(* Logix 5000 project; controller PLC_MCC1300_75F1 vendor 1 type 14 code 166 rev 32.11; software revision 32.04; part 12 of 83 *)
(* tags used below, declared in another part *)
   M302SpeedUp : MAC_SpeedUp;
   TMP_d : DINT;
   TMP_xPositioning : BOOL;
   TMP_xReverse : BOOL;
   TMP_xRun : BOOL;
   xAlwaysOFF : BOOL;
   Z300_Conveyor : UDT_StandConv[29];
   Z300_Conveyor_Conf : UDT_Conveyor_Config[29];
   Z300_Conveyor_HMW : MAC_Conveyor_ZC_HMW[29];
   Z300_Conveyor_IN_MOTION : MAC_Conveyor_ZC_IN_MOTION[29];
   Z301_HMR : MAC_Zone_ML_HMR;
(* CommandLogic, continued *)

ROUTINE M302M2_Conveyor_Output   (* ladder *)
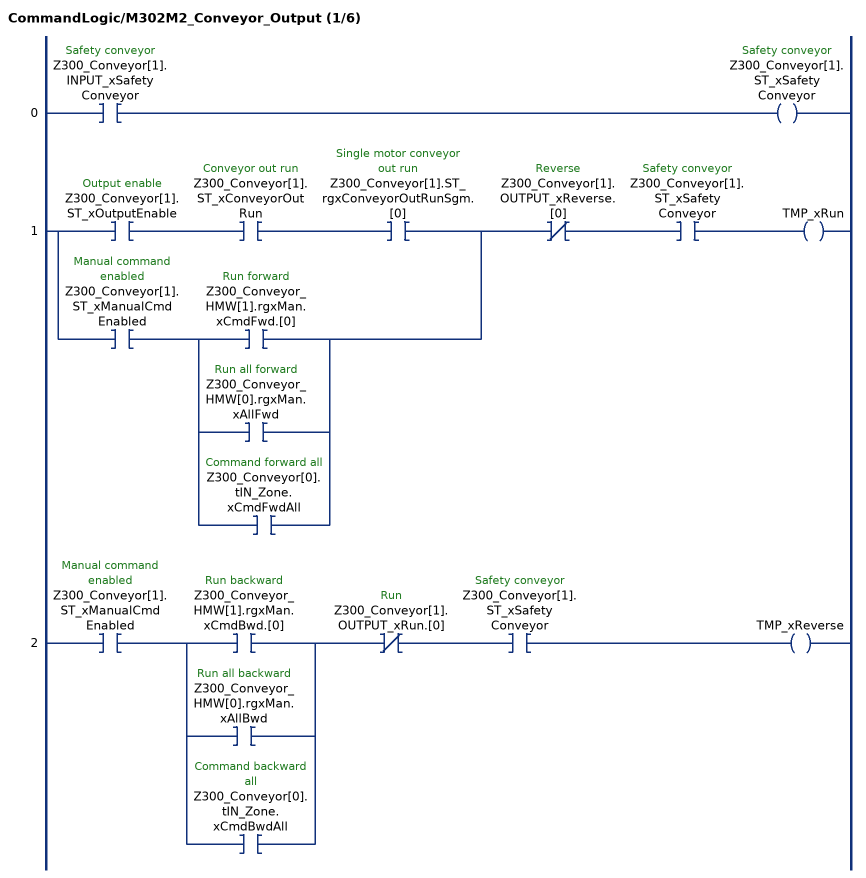
   0: XIC(Z300_Conveyor[1].INPUT_xSafetyConveyor)OTE(Z300_Conveyor[1].ST_xSafetyConveyor);
   1: [XIC(Z300_Conveyor[1].ST_xOutputEnable) XIC(Z300_Conveyor[1].ST_xConveyorOutRun) XIC(Z300_Conveyor[1].ST_rgxConveyorOutRunSgm.[0]) ,XIC(Z300_Conveyor[1].ST_xManualCmdEnabled) [XIC(Z300_Conveyor_HMW[1].rgxMan.xCmdFwd.[0]) ,XIC(Z300_Conveyor_HMW[0].rgxMan.xAllFwd) ,XIC(Z300_Conveyor[0].tIN_Zone.xCmdFwdAll) ] ]XIO(Z300_Conveyor[1].OUTPUT_xReverse.[0])XIC(Z300_Conveyor[1].ST_xSafetyConveyor)OTE(TMP_xRun);
   2: XIC(Z300_Conveyor[1].ST_xManualCmdEnabled)[XIC(Z300_Conveyor_HMW[1].rgxMan.xCmdBwd.[0]) ,XIC(Z300_Conveyor_HMW[0].rgxMan.xAllBwd) ,XIC(Z300_Conveyor[0].tIN_Zone.xCmdBwdAll) ]XIO(Z300_Conveyor[1].OUTPUT_xRun.[0])XIC(Z300_Conveyor[1].ST_xSafetyConveyor)OTE(TMP_xReverse);
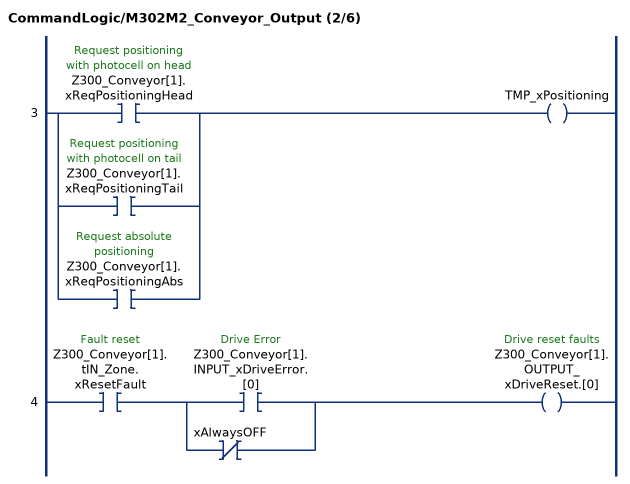
   3: [XIC(Z300_Conveyor[1].xReqPositioningHead) ,XIC(Z300_Conveyor[1].xReqPositioningTail) ,XIC(Z300_Conveyor[1].xReqPositioningAbs) ]OTE(TMP_xPositioning);
   4: XIC(Z300_Conveyor[1].tIN_Zone.xResetFault)[XIC(Z300_Conveyor[1].INPUT_xDriveError.[0]) ,XIO(xAlwaysOFF) ]OTE(Z300_Conveyor[1].OUTPUT_xDriveReset.[0]);
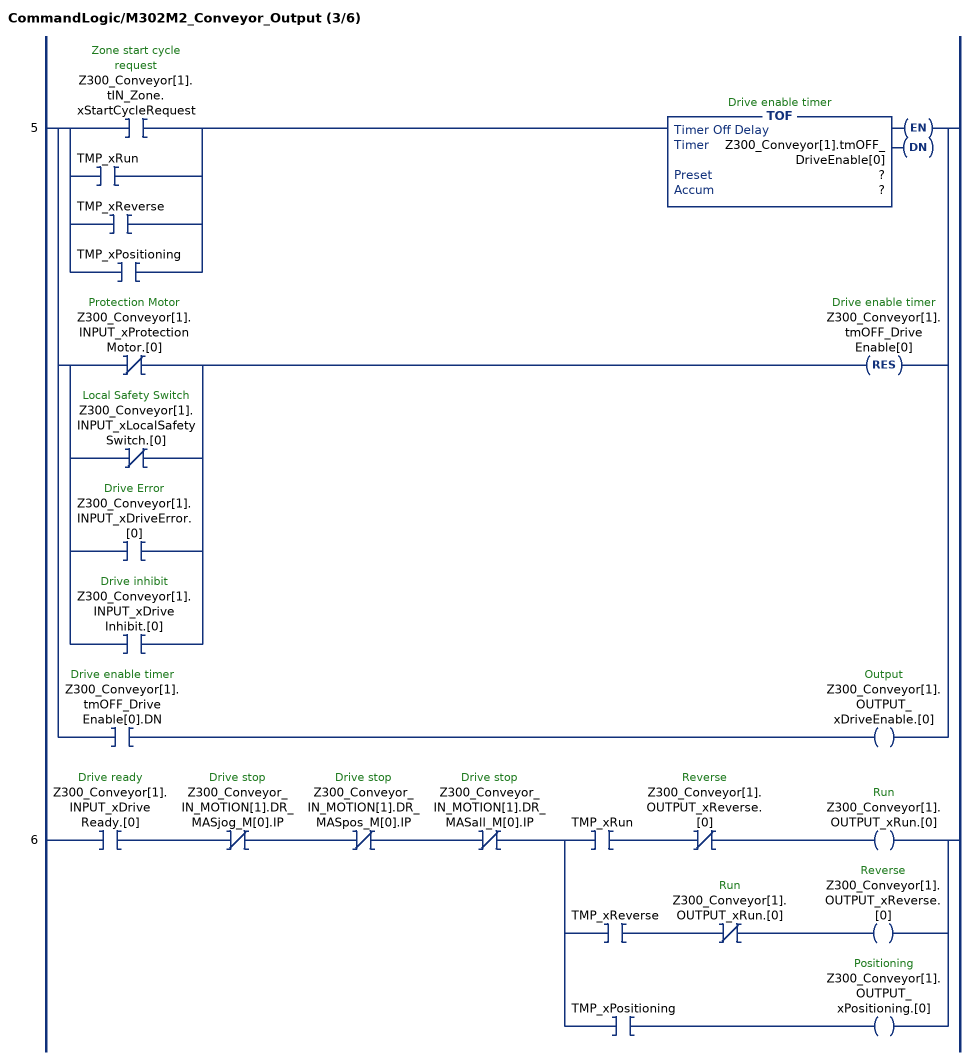
   5: [[XIC(Z300_Conveyor[1].tIN_Zone.xStartCycleRequest) ,XIC(TMP_xRun) ,XIC(TMP_xReverse) ,XIC(TMP_xPositioning) ] TOF(Z300_Conveyor[1].tmOFF_DriveEnable[0],?,?) ,[XIO(Z300_Conveyor[1].INPUT_xProtectionMotor.[0]) ,XIO(Z300_Conveyor[1].INPUT_xLocalSafetySwitch.[0]) ,XIC(Z300_Conveyor[1].INPUT_xDriveError.[0]) ,XIC(Z300_Conveyor[1].INPUT_xDriveInhibit.[0]) ] RES(Z300_Conveyor[1].tmOFF_DriveEnable[0]) ,XIC(Z300_Conveyor[1].tmOFF_DriveEnable[0].DN) OTE(Z300_Conveyor[1].OUTPUT_xDriveEnable.[0]) ];
   6: XIC(Z300_Conveyor[1].INPUT_xDriveReady.[0])XIO(Z300_Conveyor_IN_MOTION[1].DR_MASjog_M[0].IP)XIO(Z300_Conveyor_IN_MOTION[1].DR_MASpos_M[0].IP)XIO(Z300_Conveyor_IN_MOTION[1].DR_MASall_M[0].IP)[XIC(TMP_xRun) XIO(Z300_Conveyor[1].OUTPUT_xReverse.[0]) OTE(Z300_Conveyor[1].OUTPUT_xRun.[0]) ,XIC(TMP_xReverse) XIO(Z300_Conveyor[1].OUTPUT_xRun.[0]) OTE(Z300_Conveyor[1].OUTPUT_xReverse.[0]) ,XIC(TMP_xPositioning) OTE(Z300_Conveyor[1].OUTPUT_xPositioning.[0]) ];
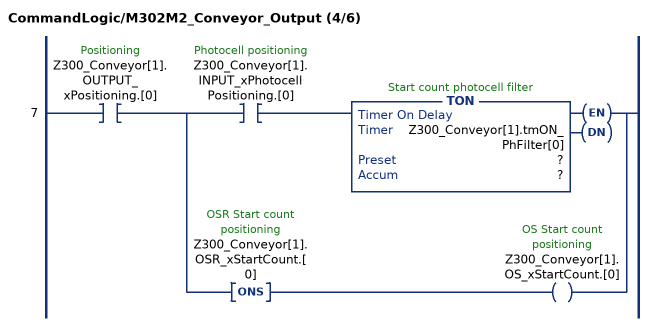
   7: XIC(Z300_Conveyor[1].OUTPUT_xPositioning.[0])[XIC(Z300_Conveyor[1].INPUT_xPhotocellPositioning.[0]) TON(Z300_Conveyor[1].tmON_PhFilter[0],?,?) ,ONS(Z300_Conveyor[1].OSR_xStartCount.[0]) OTE(Z300_Conveyor[1].OS_xStartCount.[0]) ];
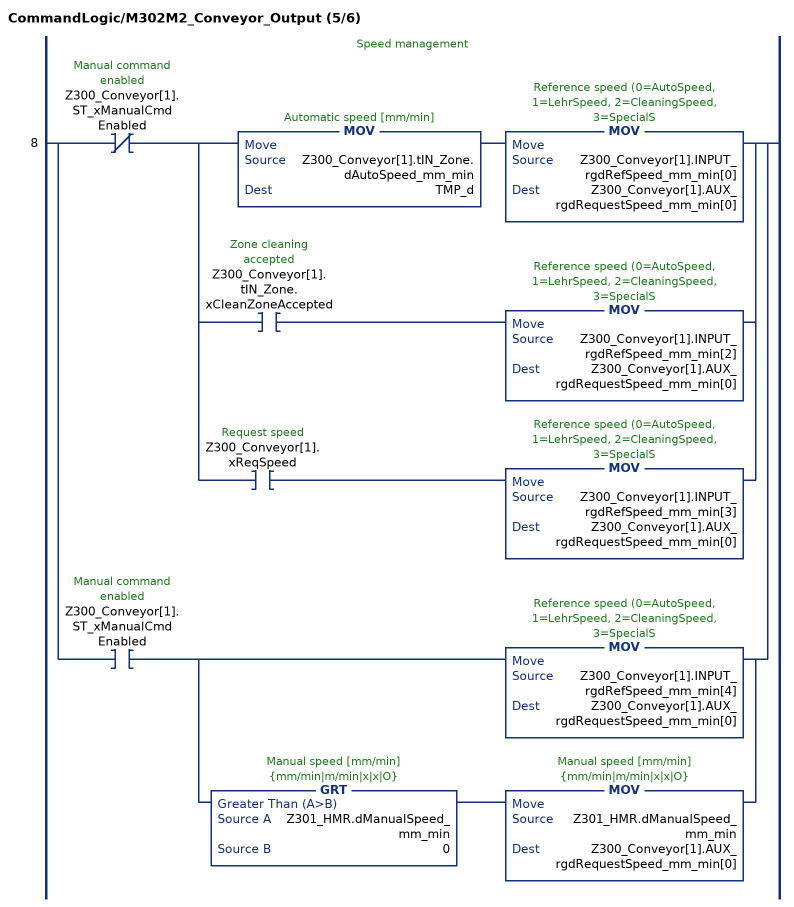
   // Speed management
   8: [XIO(Z300_Conveyor[1].ST_xManualCmdEnabled) [MOV(Z300_Conveyor[1].tIN_Zone.dAutoSpeed_mm_min,TMP_d) MOV(Z300_Conveyor[1].INPUT_rgdRefSpeed_mm_min[0],Z300_Conveyor[1].AUX_rgdRequestSpeed_mm_min[0]) ,XIC(Z300_Conveyor[1].tIN_Zone.xCleanZoneAccepted) MOV(Z300_Conveyor[1].INPUT_rgdRefSpeed_mm_min[2],Z300_Conveyor[1].AUX_rgdRequestSpeed_mm_min[0]) ,XIC(Z300_Conveyor[1].xReqSpeed) MOV(Z300_Conveyor[1].INPUT_rgdRefSpeed_mm_min[3],Z300_Conveyor[1].AUX_rgdRequestSpeed_mm_min[0]) ] ,XIC(Z300_Conveyor[1].ST_xManualCmdEnabled) [MOV(Z300_Conveyor[1].INPUT_rgdRefSpeed_mm_min[4],Z300_Conveyor[1].AUX_rgdRequestSpeed_mm_min[0]) ,GRT(Z301_HMR.dManualSpeed_mm_min,0) MOV(Z301_HMR.dManualSpeed_mm_min,Z300_Conveyor[1].AUX_rgdRequestSpeed_mm_min[0]) ] ];
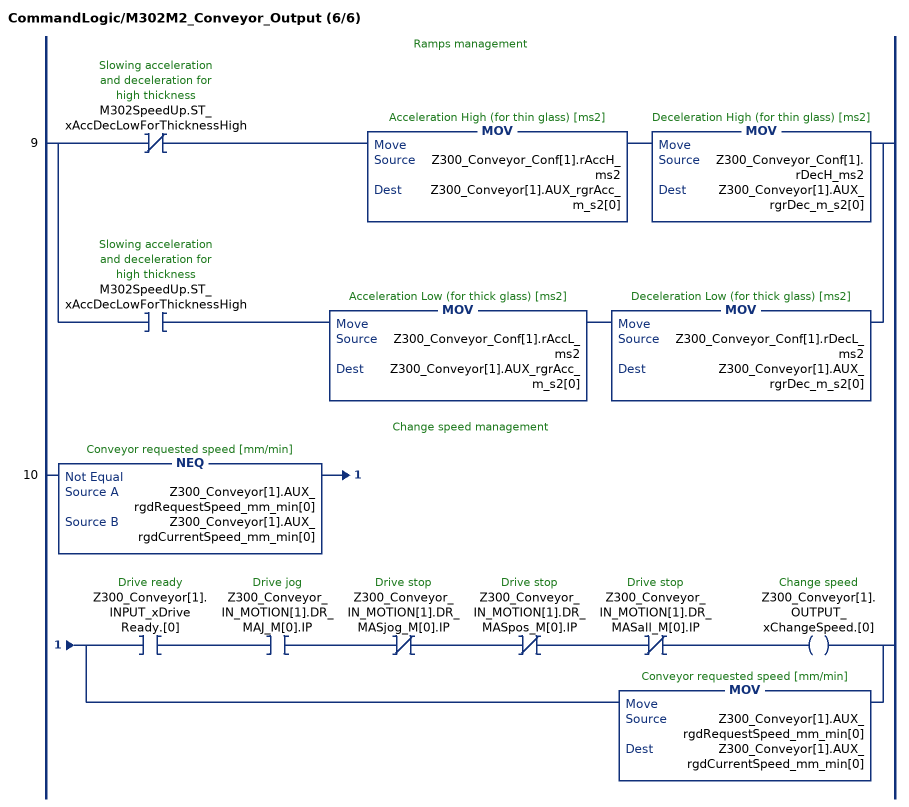
   // Ramps management
   9: [XIO(M302SpeedUp.ST_xAccDecLowForThicknessHigh) MOV(Z300_Conveyor_Conf[1].rAccH_ms2,Z300_Conveyor[1].AUX_rgrAcc_m_s2[0]) MOV(Z300_Conveyor_Conf[1].rDecH_ms2,Z300_Conveyor[1].AUX_rgrDec_m_s2[0]) ,XIC(M302SpeedUp.ST_xAccDecLowForThicknessHigh) MOV(Z300_Conveyor_Conf[1].rAccL_ms2,Z300_Conveyor[1].AUX_rgrAcc_m_s2[0]) MOV(Z300_Conveyor_Conf[1].rDecL_ms2,Z300_Conveyor[1].AUX_rgrDec_m_s2[0]) ];
   // Change speed management
   10: NEQ(Z300_Conveyor[1].AUX_rgdRequestSpeed_mm_min[0],Z300_Conveyor[1].AUX_rgdCurrentSpeed_mm_min[0])[XIC(Z300_Conveyor[1].INPUT_xDriveReady.[0]) XIC(Z300_Conveyor_IN_MOTION[1].DR_MAJ_M[0].IP) XIO(Z300_Conveyor_IN_MOTION[1].DR_MASjog_M[0].IP) XIO(Z300_Conveyor_IN_MOTION[1].DR_MASpos_M[0].IP) XIO(Z300_Conveyor_IN_MOTION[1].DR_MASall_M[0].IP) OTE(Z300_Conveyor[1].OUTPUT_xChangeSpeed.[0]) ,MOV(Z300_Conveyor[1].AUX_rgdRequestSpeed_mm_min[0],Z300_Conveyor[1].AUX_rgdCurrentSpeed_mm_min[0]) ];
END_ROUTINE

ROUTINE M302M3_Conveyor_Output   (* ladder *)
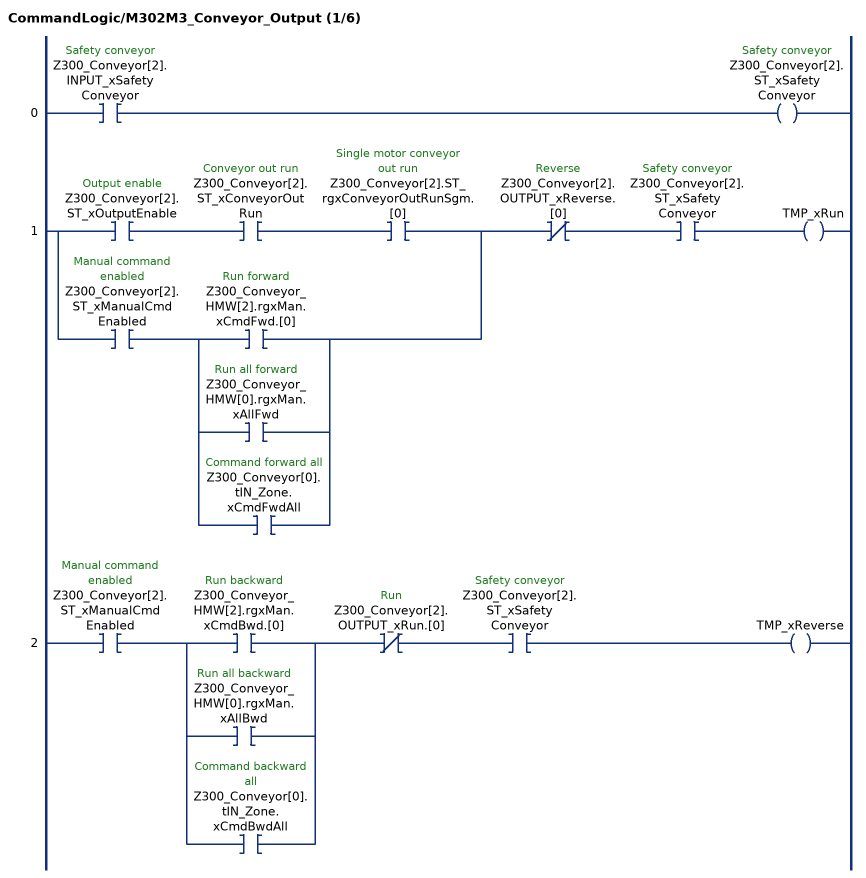
   0: XIC(Z300_Conveyor[2].INPUT_xSafetyConveyor)OTE(Z300_Conveyor[2].ST_xSafetyConveyor);
   1: [XIC(Z300_Conveyor[2].ST_xOutputEnable) XIC(Z300_Conveyor[2].ST_xConveyorOutRun) XIC(Z300_Conveyor[2].ST_rgxConveyorOutRunSgm.[0]) ,XIC(Z300_Conveyor[2].ST_xManualCmdEnabled) [XIC(Z300_Conveyor_HMW[2].rgxMan.xCmdFwd.[0]) ,XIC(Z300_Conveyor_HMW[0].rgxMan.xAllFwd) ,XIC(Z300_Conveyor[0].tIN_Zone.xCmdFwdAll) ] ]XIO(Z300_Conveyor[2].OUTPUT_xReverse.[0])XIC(Z300_Conveyor[2].ST_xSafetyConveyor)OTE(TMP_xRun);
   2: XIC(Z300_Conveyor[2].ST_xManualCmdEnabled)[XIC(Z300_Conveyor_HMW[2].rgxMan.xCmdBwd.[0]) ,XIC(Z300_Conveyor_HMW[0].rgxMan.xAllBwd) ,XIC(Z300_Conveyor[0].tIN_Zone.xCmdBwdAll) ]XIO(Z300_Conveyor[2].OUTPUT_xRun.[0])XIC(Z300_Conveyor[2].ST_xSafetyConveyor)OTE(TMP_xReverse);
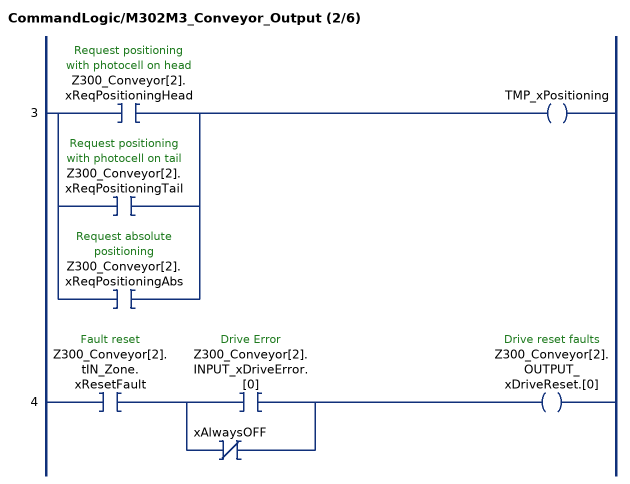
   3: [XIC(Z300_Conveyor[2].xReqPositioningHead) ,XIC(Z300_Conveyor[2].xReqPositioningTail) ,XIC(Z300_Conveyor[2].xReqPositioningAbs) ]OTE(TMP_xPositioning);
   4: XIC(Z300_Conveyor[2].tIN_Zone.xResetFault)[XIC(Z300_Conveyor[2].INPUT_xDriveError.[0]) ,XIO(xAlwaysOFF) ]OTE(Z300_Conveyor[2].OUTPUT_xDriveReset.[0]);
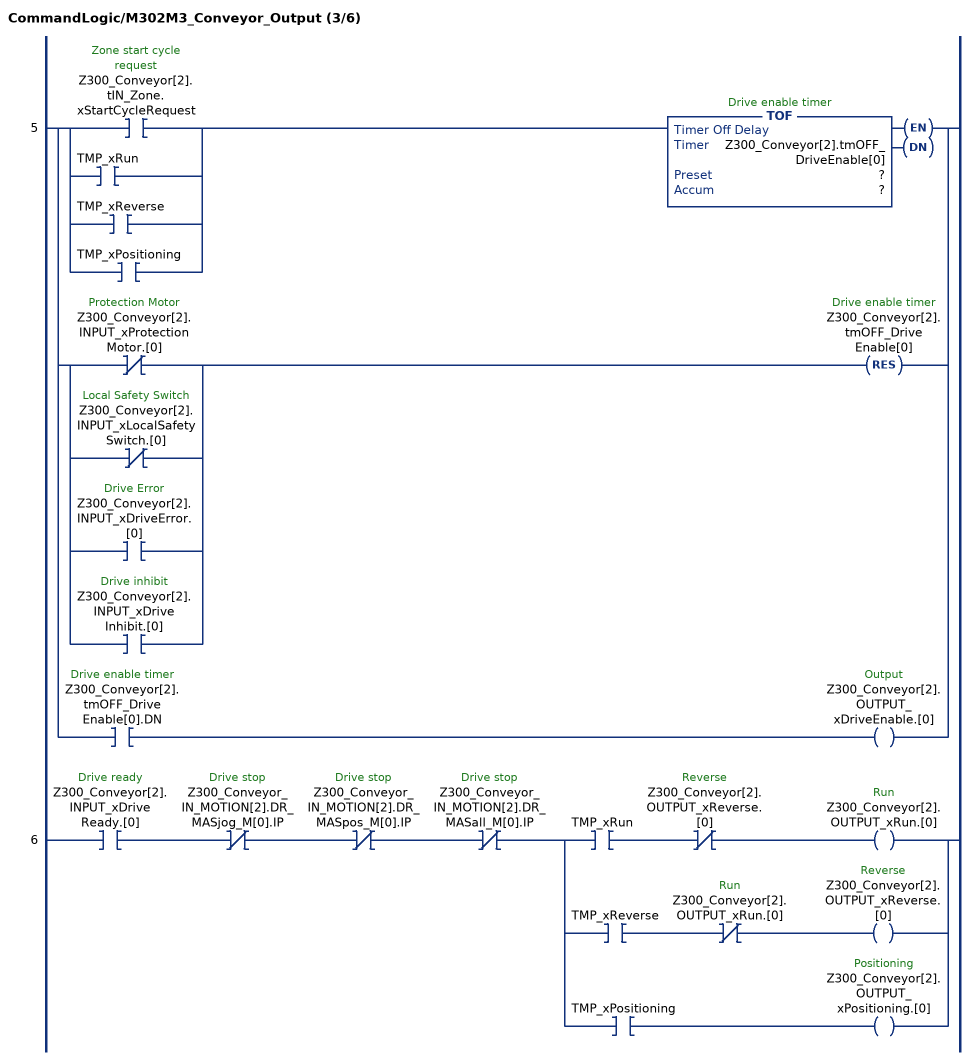
   5: [[XIC(Z300_Conveyor[2].tIN_Zone.xStartCycleRequest) ,XIC(TMP_xRun) ,XIC(TMP_xReverse) ,XIC(TMP_xPositioning) ] TOF(Z300_Conveyor[2].tmOFF_DriveEnable[0],?,?) ,[XIO(Z300_Conveyor[2].INPUT_xProtectionMotor.[0]) ,XIO(Z300_Conveyor[2].INPUT_xLocalSafetySwitch.[0]) ,XIC(Z300_Conveyor[2].INPUT_xDriveError.[0]) ,XIC(Z300_Conveyor[2].INPUT_xDriveInhibit.[0]) ] RES(Z300_Conveyor[2].tmOFF_DriveEnable[0]) ,XIC(Z300_Conveyor[2].tmOFF_DriveEnable[0].DN) OTE(Z300_Conveyor[2].OUTPUT_xDriveEnable.[0]) ];
   6: XIC(Z300_Conveyor[2].INPUT_xDriveReady.[0])XIO(Z300_Conveyor_IN_MOTION[2].DR_MASjog_M[0].IP)XIO(Z300_Conveyor_IN_MOTION[2].DR_MASpos_M[0].IP)XIO(Z300_Conveyor_IN_MOTION[2].DR_MASall_M[0].IP)[XIC(TMP_xRun) XIO(Z300_Conveyor[2].OUTPUT_xReverse.[0]) OTE(Z300_Conveyor[2].OUTPUT_xRun.[0]) ,XIC(TMP_xReverse) XIO(Z300_Conveyor[2].OUTPUT_xRun.[0]) OTE(Z300_Conveyor[2].OUTPUT_xReverse.[0]) ,XIC(TMP_xPositioning) OTE(Z300_Conveyor[2].OUTPUT_xPositioning.[0]) ];
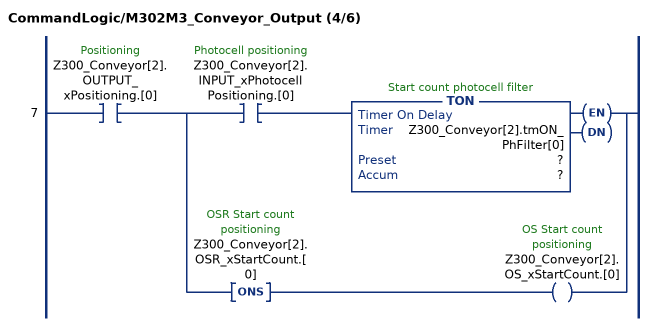
   7: XIC(Z300_Conveyor[2].OUTPUT_xPositioning.[0])[XIC(Z300_Conveyor[2].INPUT_xPhotocellPositioning.[0]) TON(Z300_Conveyor[2].tmON_PhFilter[0],?,?) ,ONS(Z300_Conveyor[2].OSR_xStartCount.[0]) OTE(Z300_Conveyor[2].OS_xStartCount.[0]) ];
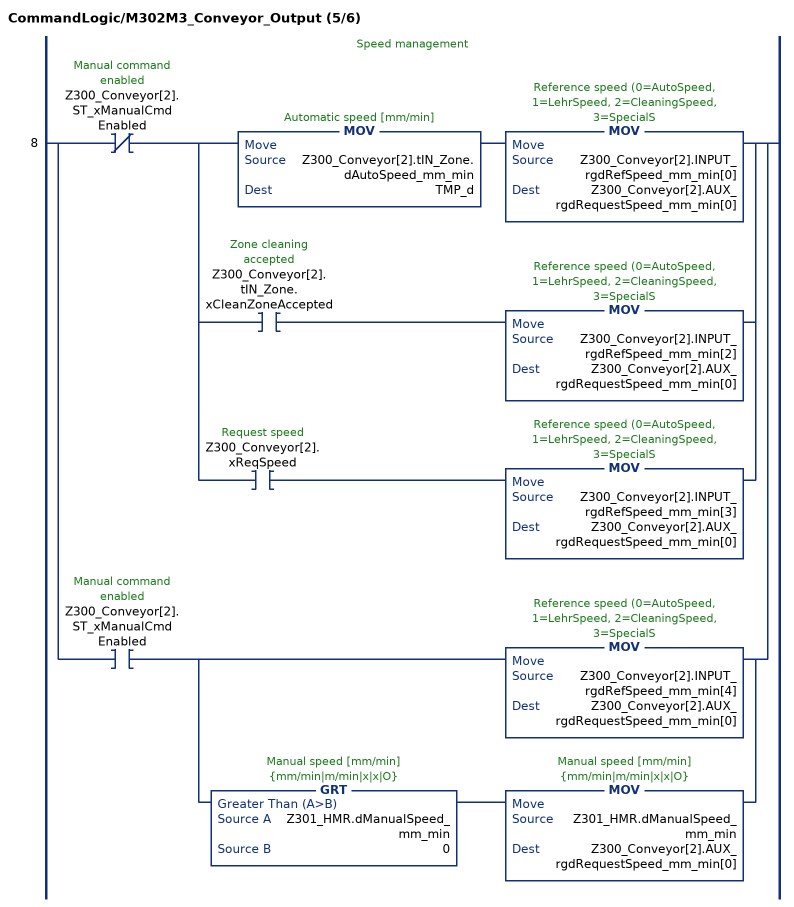
   // Speed management
   8: [XIO(Z300_Conveyor[2].ST_xManualCmdEnabled) [MOV(Z300_Conveyor[2].tIN_Zone.dAutoSpeed_mm_min,TMP_d) MOV(Z300_Conveyor[2].INPUT_rgdRefSpeed_mm_min[0],Z300_Conveyor[2].AUX_rgdRequestSpeed_mm_min[0]) ,XIC(Z300_Conveyor[2].tIN_Zone.xCleanZoneAccepted) MOV(Z300_Conveyor[2].INPUT_rgdRefSpeed_mm_min[2],Z300_Conveyor[2].AUX_rgdRequestSpeed_mm_min[0]) ,XIC(Z300_Conveyor[2].xReqSpeed) MOV(Z300_Conveyor[2].INPUT_rgdRefSpeed_mm_min[3],Z300_Conveyor[2].AUX_rgdRequestSpeed_mm_min[0]) ] ,XIC(Z300_Conveyor[2].ST_xManualCmdEnabled) [MOV(Z300_Conveyor[2].INPUT_rgdRefSpeed_mm_min[4],Z300_Conveyor[2].AUX_rgdRequestSpeed_mm_min[0]) ,GRT(Z301_HMR.dManualSpeed_mm_min,0) MOV(Z301_HMR.dManualSpeed_mm_min,Z300_Conveyor[2].AUX_rgdRequestSpeed_mm_min[0]) ] ];
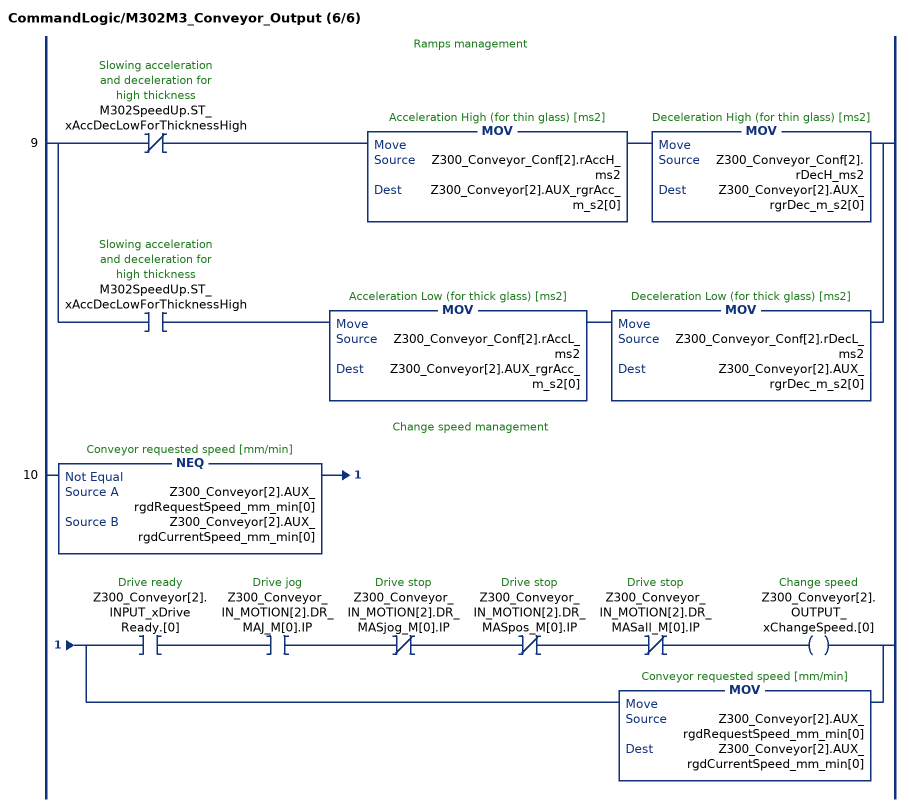
   // Ramps management
   9: [XIO(M302SpeedUp.ST_xAccDecLowForThicknessHigh) MOV(Z300_Conveyor_Conf[2].rAccH_ms2,Z300_Conveyor[2].AUX_rgrAcc_m_s2[0]) MOV(Z300_Conveyor_Conf[2].rDecH_ms2,Z300_Conveyor[2].AUX_rgrDec_m_s2[0]) ,XIC(M302SpeedUp.ST_xAccDecLowForThicknessHigh) MOV(Z300_Conveyor_Conf[2].rAccL_ms2,Z300_Conveyor[2].AUX_rgrAcc_m_s2[0]) MOV(Z300_Conveyor_Conf[2].rDecL_ms2,Z300_Conveyor[2].AUX_rgrDec_m_s2[0]) ];
   // Change speed management
   10: NEQ(Z300_Conveyor[2].AUX_rgdRequestSpeed_mm_min[0],Z300_Conveyor[2].AUX_rgdCurrentSpeed_mm_min[0])[XIC(Z300_Conveyor[2].INPUT_xDriveReady.[0]) XIC(Z300_Conveyor_IN_MOTION[2].DR_MAJ_M[0].IP) XIO(Z300_Conveyor_IN_MOTION[2].DR_MASjog_M[0].IP) XIO(Z300_Conveyor_IN_MOTION[2].DR_MASpos_M[0].IP) XIO(Z300_Conveyor_IN_MOTION[2].DR_MASall_M[0].IP) OTE(Z300_Conveyor[2].OUTPUT_xChangeSpeed.[0]) ,MOV(Z300_Conveyor[2].AUX_rgdRequestSpeed_mm_min[0],Z300_Conveyor[2].AUX_rgdCurrentSpeed_mm_min[0]) ];
END_ROUTINE

ROUTINE M302M4_Conveyor_Output   (* ladder *)
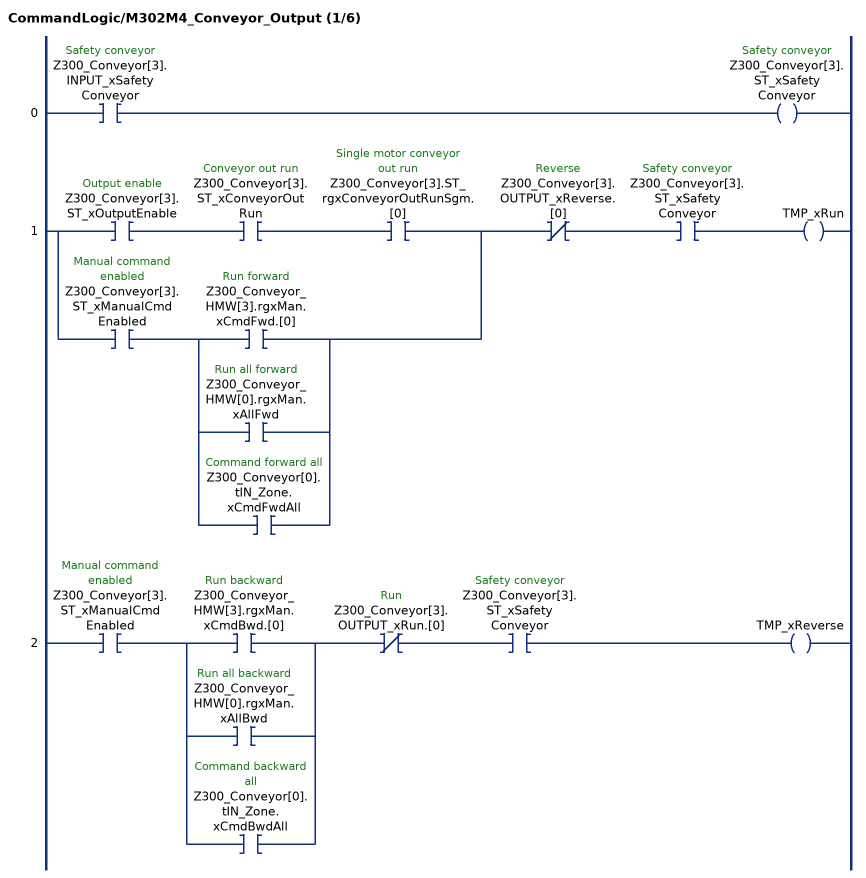
   0: XIC(Z300_Conveyor[3].INPUT_xSafetyConveyor)OTE(Z300_Conveyor[3].ST_xSafetyConveyor);
   1: [XIC(Z300_Conveyor[3].ST_xOutputEnable) XIC(Z300_Conveyor[3].ST_xConveyorOutRun) XIC(Z300_Conveyor[3].ST_rgxConveyorOutRunSgm.[0]) ,XIC(Z300_Conveyor[3].ST_xManualCmdEnabled) [XIC(Z300_Conveyor_HMW[3].rgxMan.xCmdFwd.[0]) ,XIC(Z300_Conveyor_HMW[0].rgxMan.xAllFwd) ,XIC(Z300_Conveyor[0].tIN_Zone.xCmdFwdAll) ] ]XIO(Z300_Conveyor[3].OUTPUT_xReverse.[0])XIC(Z300_Conveyor[3].ST_xSafetyConveyor)OTE(TMP_xRun);
   2: XIC(Z300_Conveyor[3].ST_xManualCmdEnabled)[XIC(Z300_Conveyor_HMW[3].rgxMan.xCmdBwd.[0]) ,XIC(Z300_Conveyor_HMW[0].rgxMan.xAllBwd) ,XIC(Z300_Conveyor[0].tIN_Zone.xCmdBwdAll) ]XIO(Z300_Conveyor[3].OUTPUT_xRun.[0])XIC(Z300_Conveyor[3].ST_xSafetyConveyor)OTE(TMP_xReverse);
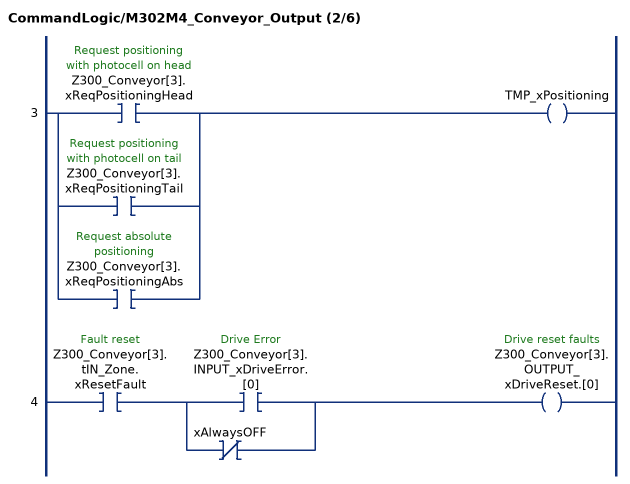
   3: [XIC(Z300_Conveyor[3].xReqPositioningHead) ,XIC(Z300_Conveyor[3].xReqPositioningTail) ,XIC(Z300_Conveyor[3].xReqPositioningAbs) ]OTE(TMP_xPositioning);
   4: XIC(Z300_Conveyor[3].tIN_Zone.xResetFault)[XIC(Z300_Conveyor[3].INPUT_xDriveError.[0]) ,XIO(xAlwaysOFF) ]OTE(Z300_Conveyor[3].OUTPUT_xDriveReset.[0]);
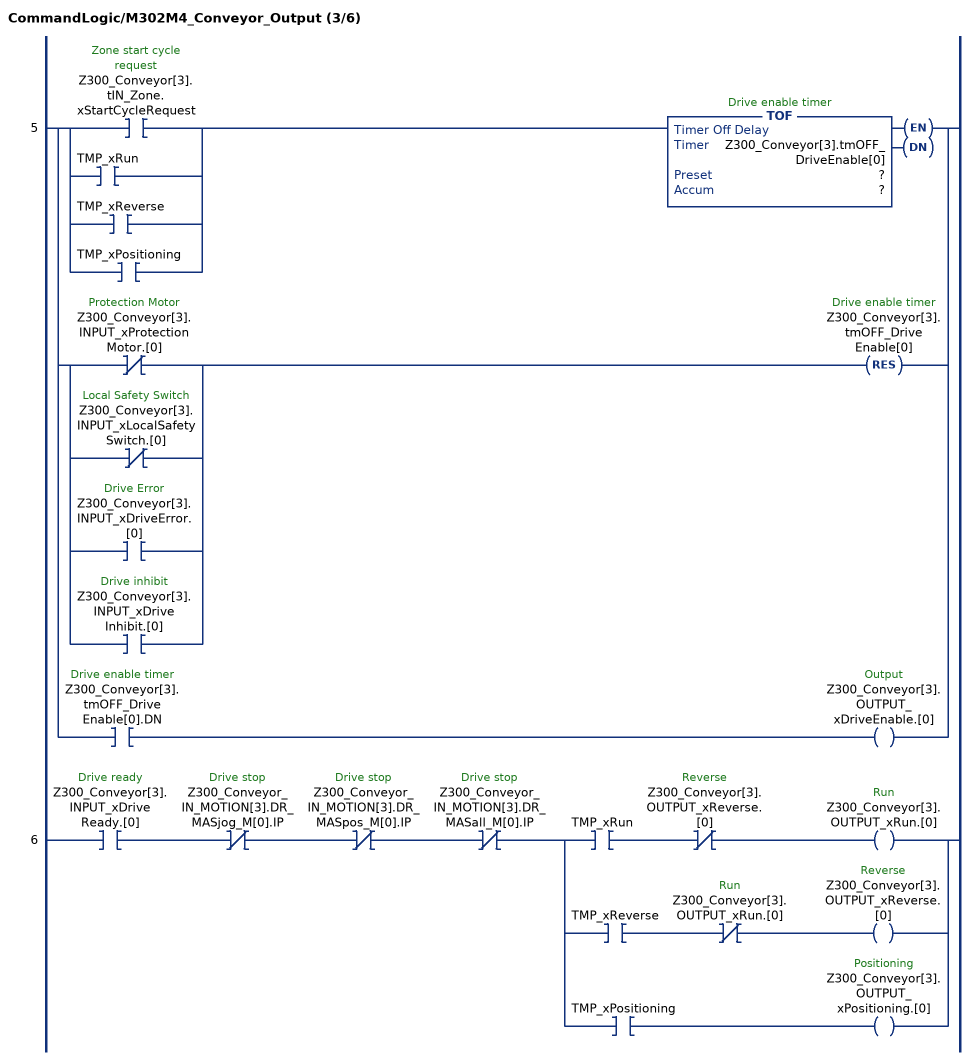
   5: [[XIC(Z300_Conveyor[3].tIN_Zone.xStartCycleRequest) ,XIC(TMP_xRun) ,XIC(TMP_xReverse) ,XIC(TMP_xPositioning) ] TOF(Z300_Conveyor[3].tmOFF_DriveEnable[0],?,?) ,[XIO(Z300_Conveyor[3].INPUT_xProtectionMotor.[0]) ,XIO(Z300_Conveyor[3].INPUT_xLocalSafetySwitch.[0]) ,XIC(Z300_Conveyor[3].INPUT_xDriveError.[0]) ,XIC(Z300_Conveyor[3].INPUT_xDriveInhibit.[0]) ] RES(Z300_Conveyor[3].tmOFF_DriveEnable[0]) ,XIC(Z300_Conveyor[3].tmOFF_DriveEnable[0].DN) OTE(Z300_Conveyor[3].OUTPUT_xDriveEnable.[0]) ];
   6: XIC(Z300_Conveyor[3].INPUT_xDriveReady.[0])XIO(Z300_Conveyor_IN_MOTION[3].DR_MASjog_M[0].IP)XIO(Z300_Conveyor_IN_MOTION[3].DR_MASpos_M[0].IP)XIO(Z300_Conveyor_IN_MOTION[3].DR_MASall_M[0].IP)[XIC(TMP_xRun) XIO(Z300_Conveyor[3].OUTPUT_xReverse.[0]) OTE(Z300_Conveyor[3].OUTPUT_xRun.[0]) ,XIC(TMP_xReverse) XIO(Z300_Conveyor[3].OUTPUT_xRun.[0]) OTE(Z300_Conveyor[3].OUTPUT_xReverse.[0]) ,XIC(TMP_xPositioning) OTE(Z300_Conveyor[3].OUTPUT_xPositioning.[0]) ];
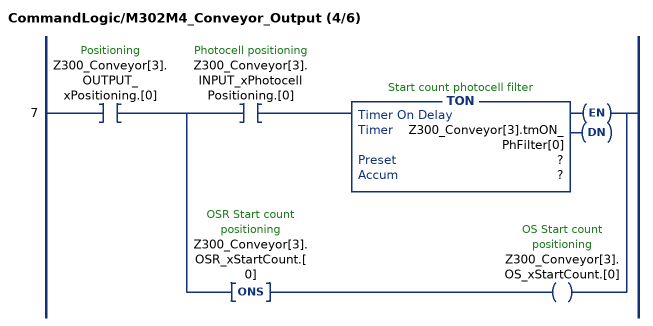
   7: XIC(Z300_Conveyor[3].OUTPUT_xPositioning.[0])[XIC(Z300_Conveyor[3].INPUT_xPhotocellPositioning.[0]) TON(Z300_Conveyor[3].tmON_PhFilter[0],?,?) ,ONS(Z300_Conveyor[3].OSR_xStartCount.[0]) OTE(Z300_Conveyor[3].OS_xStartCount.[0]) ];
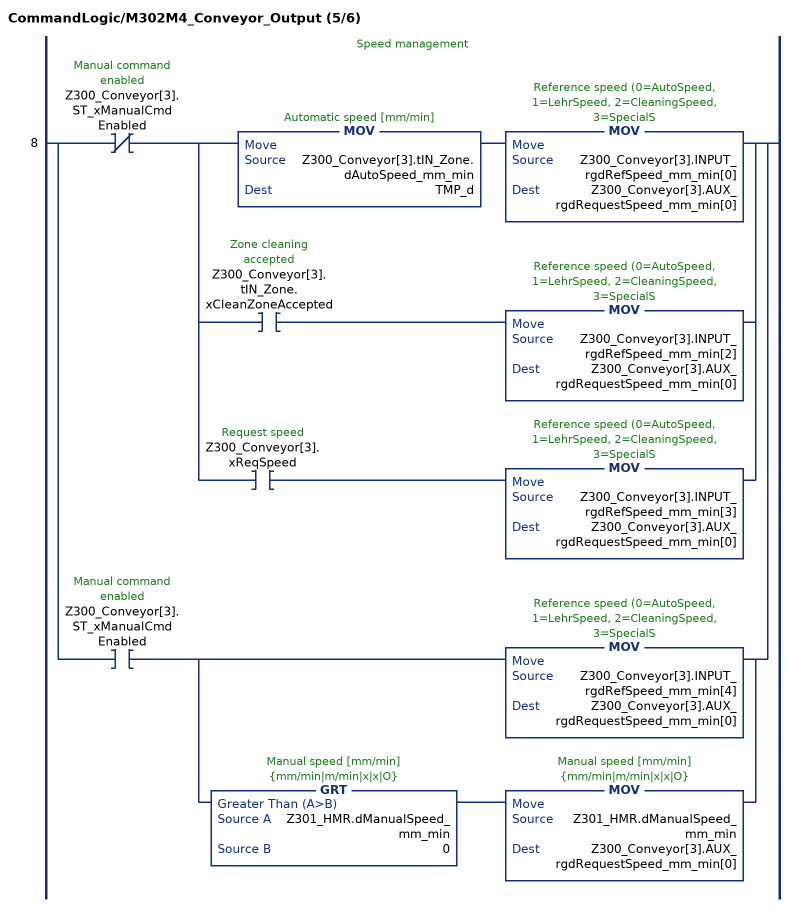
   // Speed management
   8: [XIO(Z300_Conveyor[3].ST_xManualCmdEnabled) [MOV(Z300_Conveyor[3].tIN_Zone.dAutoSpeed_mm_min,TMP_d) MOV(Z300_Conveyor[3].INPUT_rgdRefSpeed_mm_min[0],Z300_Conveyor[3].AUX_rgdRequestSpeed_mm_min[0]) ,XIC(Z300_Conveyor[3].tIN_Zone.xCleanZoneAccepted) MOV(Z300_Conveyor[3].INPUT_rgdRefSpeed_mm_min[2],Z300_Conveyor[3].AUX_rgdRequestSpeed_mm_min[0]) ,XIC(Z300_Conveyor[3].xReqSpeed) MOV(Z300_Conveyor[3].INPUT_rgdRefSpeed_mm_min[3],Z300_Conveyor[3].AUX_rgdRequestSpeed_mm_min[0]) ] ,XIC(Z300_Conveyor[3].ST_xManualCmdEnabled) [MOV(Z300_Conveyor[3].INPUT_rgdRefSpeed_mm_min[4],Z300_Conveyor[3].AUX_rgdRequestSpeed_mm_min[0]) ,GRT(Z301_HMR.dManualSpeed_mm_min,0) MOV(Z301_HMR.dManualSpeed_mm_min,Z300_Conveyor[3].AUX_rgdRequestSpeed_mm_min[0]) ] ];
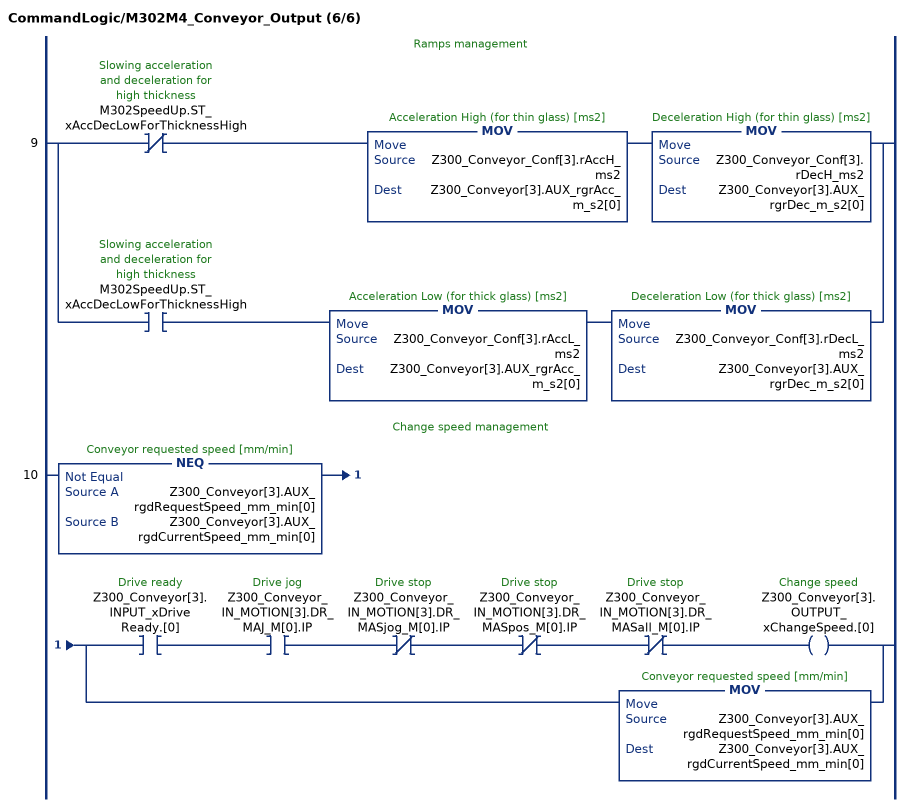
   // Ramps management
   9: [XIO(M302SpeedUp.ST_xAccDecLowForThicknessHigh) MOV(Z300_Conveyor_Conf[3].rAccH_ms2,Z300_Conveyor[3].AUX_rgrAcc_m_s2[0]) MOV(Z300_Conveyor_Conf[3].rDecH_ms2,Z300_Conveyor[3].AUX_rgrDec_m_s2[0]) ,XIC(M302SpeedUp.ST_xAccDecLowForThicknessHigh) MOV(Z300_Conveyor_Conf[3].rAccL_ms2,Z300_Conveyor[3].AUX_rgrAcc_m_s2[0]) MOV(Z300_Conveyor_Conf[3].rDecL_ms2,Z300_Conveyor[3].AUX_rgrDec_m_s2[0]) ];
   // Change speed management
   10: NEQ(Z300_Conveyor[3].AUX_rgdRequestSpeed_mm_min[0],Z300_Conveyor[3].AUX_rgdCurrentSpeed_mm_min[0])[XIC(Z300_Conveyor[3].INPUT_xDriveReady.[0]) XIC(Z300_Conveyor_IN_MOTION[3].DR_MAJ_M[0].IP) XIO(Z300_Conveyor_IN_MOTION[3].DR_MASjog_M[0].IP) XIO(Z300_Conveyor_IN_MOTION[3].DR_MASpos_M[0].IP) XIO(Z300_Conveyor_IN_MOTION[3].DR_MASall_M[0].IP) OTE(Z300_Conveyor[3].OUTPUT_xChangeSpeed.[0]) ,MOV(Z300_Conveyor[3].AUX_rgdRequestSpeed_mm_min[0],Z300_Conveyor[3].AUX_rgdCurrentSpeed_mm_min[0]) ];
END_ROUTINE
